REGION Network 3: Ya buscó caja DESACTIVADO
   // Detecta cuando el brazo de succion se encuentra arriba y setea una marca "ya buscó caja". La cinta no va a arrancar hasta que esta marca YA BUSCO CAJA se active.
   RUNG wire#powerrail
      Contact( "Marcha" )
      Contact( "iSNS_bs_arriba" )
      I_Contact( "iSNS_bs_abajo" )
      S_SR(operand := "Aux1", r1 := wire#w1)
      Coil( "Ya buscó caja" )
   END_RUNG
   RUNG wire#powerrail
      I_Contact( "Marcha" )
   END_RUNG wire#w1
   RUNG wire#powerrail
      { S7_Templates := "SrcType := DInt" } GE_Contact(in1 := "Encoder", in2 := 20)
      { S7_Templates := "SrcType := DInt" } LT_Contact(in1 := "Encoder", in2 := 45)
   END_RUNG wire#w1
   RUNG wire#powerrail
      Contact( "Habilita modo Probar" )
   END_RUNG wire#w1
   // the same network as SCL:
   IF "Marcha" AND "iSNS_bs_arriba" AND NOT "iSNS_bs_abajo" THEN
       "Aux1" := TRUE;   // SR flip-flop
   END_IF;
   IF NOT "Marcha" OR (("Encoder" >= 20) AND ("Encoder" < 45)) OR "Habilita modo Probar" THEN
       "Aux1" := FALSE;
   END_IF;
   "Ya buscó caja" := "Aux1";
END_REGION

REGION Network 4: Activa los succionadores.
   "TOFF".TOF(IN := NOT "iSNS_bs_abajo", PT := T#300ms);
   "Activa succionadores" := "TOFF".Q;
END_REGION

REGION Network 5: Cuando el brazo llega hasta abajo, lo detiene por 300 ms para asegurar que la caja salió de su rango. DESACTIVADO
   // DESACTIVADO
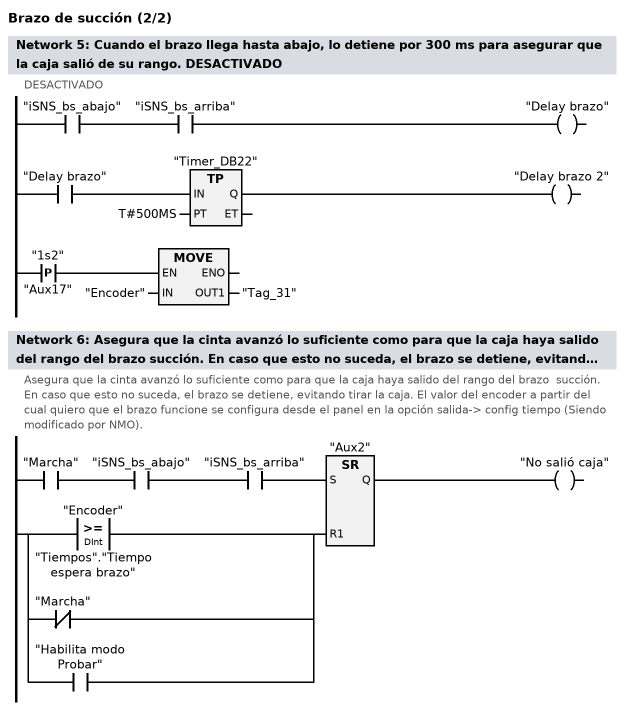
   "Delay brazo" := "iSNS_bs_abajo" AND "iSNS_bs_arriba";
   "Timer_DB22".TP(IN := "Delay brazo", PT := T#500MS);
   "Delay brazo 2" := "Timer_DB22".Q;
   #_w1 := "1s2" AND NOT "Aux17";   // rising edge of "1s2"
   "Aux17" := "1s2";
   IF #_w1 THEN "Tag_31" := "Encoder"; END_IF;
END_REGION

REGION Network 6: Asegura que la cinta avanzó lo suficiente como para que la caja haya salido del rango del brazo succión. En caso que esto no suceda, el brazo se detiene, evitando tirar la caja
   // Asegura que la cinta avanzó lo suficiente como para que la caja haya salido del rango del brazo  succión. En caso que esto no suceda, el brazo se detiene, evitando tirar la caja. El valor del encoder a partir del cual quiero que el brazo funcione se configura desde el panel en la opción salida-> config tiempo (Siendo modificado por NMO).
   RUNG wire#powerrail
      Contact( "Marcha" )
      Contact( "iSNS_bs_abajo" )
      Contact( "iSNS_bs_arriba" )
      S_SR(operand := "Aux2", r1 := wire#w1)
      Coil( "No salió caja" )
   END_RUNG
   RUNG wire#powerrail
      { S7_Templates := "SrcType := DInt" } GE_Contact(in1 := "Encoder", in2 := "Tiempos"."Tiempo espera brazo")
   END_RUNG wire#w1
   RUNG wire#powerrail
      I_Contact( "Marcha" )
   END_RUNG wire#w1
   RUNG wire#powerrail
      Contact( "Habilita modo Probar" )
   END_RUNG wire#w1
   // the same network as SCL:
   IF "Marcha" AND "iSNS_bs_abajo" AND "iSNS_bs_arriba" THEN
       "Aux2" := TRUE;   // SR flip-flop
   END_IF;
   IF ("Encoder" >= "Tiempos"."Tiempo espera brazo") OR NOT "Marcha" OR "Habilita modo Probar" THEN
       "Aux2" := FALSE;
   END_IF;
   "No salió caja" := "Aux2";
END_REGION
END_FUNCTION

ORGANIZATION_BLOCK "Main"   // OB1, LAD, ProgramCycle
TITLE = "Main Program Sweep (Cycle)"
{ S7_Optimized_Access := 'TRUE' }
VERSION : 0.1
BEGIN

REGION Network 1: Inversión de algunas entradas
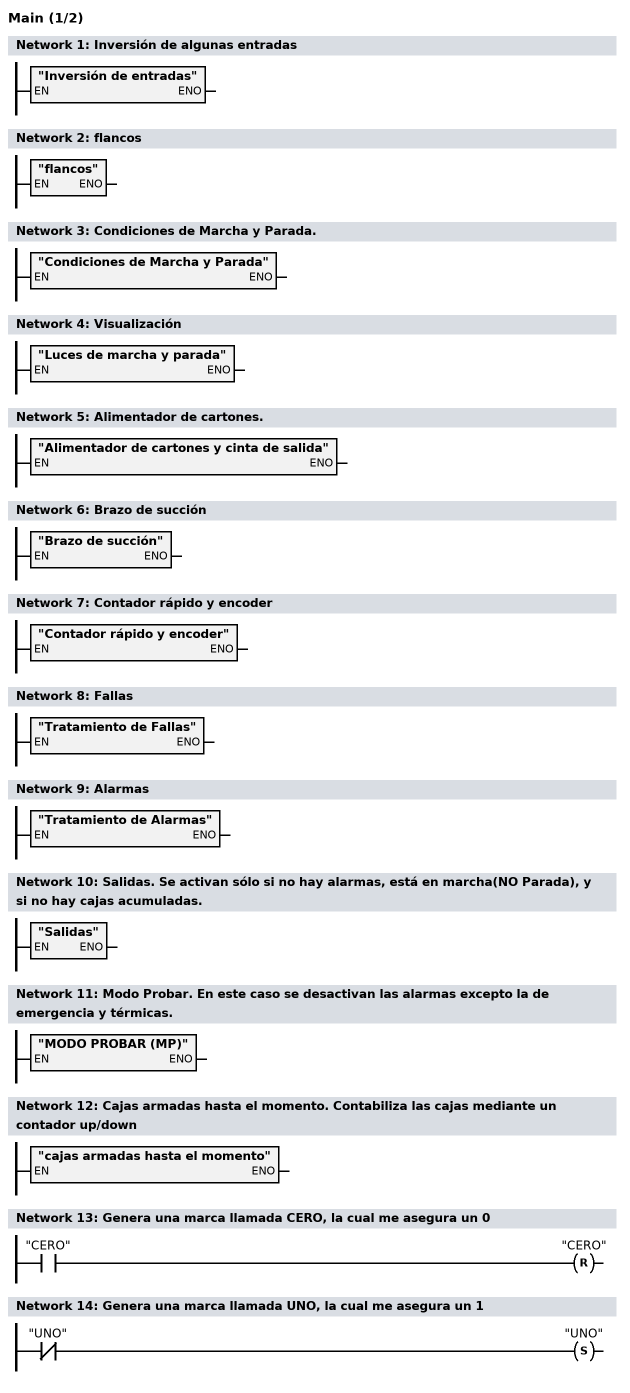
   RUNG wire#powerrail
      "Inversión de entradas"()
   END_RUNG
   // the same network as SCL:
   "Inversión de entradas"();
END_REGION

REGION Network 2: flancos
   RUNG wire#powerrail
      "flancos"()
   END_RUNG
   // the same network as SCL:
   "flancos"();
END_REGION

REGION Network 3: Condiciones de Marcha y Parada.
   RUNG wire#powerrail
      "Condiciones de Marcha y Parada"()
   END_RUNG
   // the same network as SCL:
   "Condiciones de Marcha y Parada"();
END_REGION

REGION Network 4: Visualización
   RUNG wire#powerrail
      "Luces de marcha y parada"()
   END_RUNG
   // the same network as SCL:
   "Luces de marcha y parada"();
END_REGION

REGION Network 5: Alimentador de cartones.
   RUNG wire#powerrail
      "Alimentador de cartones y cinta de salida"()
   END_RUNG
   // the same network as SCL:
   "Alimentador de cartones y cinta de salida"();
END_REGION

REGION Network 6: Brazo de succión
   RUNG wire#powerrail
      "Brazo de succión"()
   END_RUNG
   // the same network as SCL:
   "Brazo de succión"();
END_REGION

REGION Network 7: Contador rápido y encoder
   RUNG wire#powerrail
      "Contador rápido y encoder"()
   END_RUNG
   // the same network as SCL:
   "Contador rápido y encoder"();
END_REGION

REGION Network 8: Fallas
   RUNG wire#powerrail
      "Tratamiento de Fallas"()
   END_RUNG
   // the same network as SCL:
   "Tratamiento de Fallas"();
END_REGION

REGION Network 9: Alarmas
   RUNG wire#powerrail
      "Tratamiento de Alarmas"()
   END_RUNG
   // the same network as SCL:
   "Tratamiento de Alarmas"();
END_REGION

REGION Network 10: Salidas. Se activan sólo si no hay alarmas, está en marcha(NO Parada), y si no hay cajas acumuladas.
   RUNG wire#powerrail
      "Salidas"()
   END_RUNG
   // the same network as SCL:
   "Salidas"();
END_REGION

REGION Network 11: Modo Probar. En este caso se desactivan las alarmas excepto la de emergencia y térmicas.
   RUNG wire#powerrail
      "MODO PROBAR (MP)"()
   END_RUNG
   // the same network as SCL:
   "MODO PROBAR (MP)"();
END_REGION

REGION Network 12: Cajas armadas hasta el momento. Contabiliza las cajas mediante un contador up/down
   RUNG wire#powerrail
      "cajas armadas hasta el momento"()
   END_RUNG
   // the same network as SCL:
   "cajas armadas hasta el momento"();
END_REGION

REGION Network 13: Genera una marca llamada CERO, la cual me asegura un 0
   RUNG wire#powerrail
      Contact( "CERO" )
      R_Coil( "CERO" )
   END_RUNG
   // the same network as SCL:
   IF "CERO" THEN "CERO" := FALSE; END_IF;
END_REGION

REGION Network 14: Genera una marca llamada UNO, la cual me asegura un 1
   RUNG wire#powerrail
      I_Contact( "UNO" )
      S_Coil( "UNO" )
   END_RUNG
   // the same network as SCL:
   IF NOT "UNO" THEN "UNO" := TRUE; END_IF;
END_REGION

REGION Network 15: Secuencia Principal
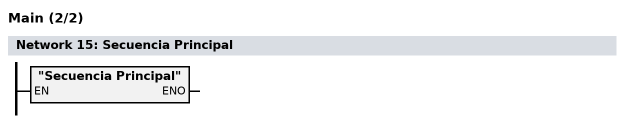
   RUNG wire#powerrail
      "Secuencia Principal"()
   END_RUNG
   // the same network as SCL:
   "Secuencia Principal"();
END_REGION
END_ORGANIZATION_BLOCK

(* ===== HMI "HMI_RT_1" =====
system functions are stored by id; their names below are inferred from use
connection "Conexión_HMI": ETHERNET, SMART_S7_1200_OMS

HMI tags "Tabla de variables estándar"
   "Alarmas_1" : Word AT %DB19.DBW0, 1 s
   "Alarmas_2" : Word AT %DB19.DBW2, 1 s
   "iAveria-reposicion" : Bool = PLC "iAveria-reposicion" AT %I32.2, 1 s
   "olmpR" : Bool = PLC oLmpR AT %Q32.5, 1 s
   "serie de fallas" : Bool = PLC "Serie de fallas" AT %M24.7, 1 s
   "Rearme desde panel" : Bool = PLC "Rearme desde panel" AT %M25.0, 1 s
   "olmpV" : Bool = PLC oLmpV AT %Q32.6, 1 s
   "SNS_carton en area de colado" : Bool = PLC "iSNS_carton en area de colado" AT %I33.3, 1 s
   "SNS_bs_arriba" : Bool = PLC iSNS_bs_arriba AT %I33.7, 1 s
   "SNS_bs_abajo" : Bool = PLC iSNS_bs_abajo AT %I33.6, 1 s
   "sns_nivel_bajo_cartones" : Bool = PLC iSNS_nivel_bajo_cartones AT %I33.0, 1 s
   "SNSpush_atras" : Bool = PLC iSNSpush_atras AT %I33.2, 1 s
   "SNSpush_adel" : Bool = PLC iSNSpush_adel AT %I0.2, 1 s
   "SNSpegamento en depósito" : Bool = PLC "iSNSpegamento en depósito" AT %I1.2, 1 s
   "SNScaja_trab" : Bool = PLC iSNScaja_trab AT %I1.4, 1 s
   "SNSalp" : Bool = PLC iSNSalp AT %I1.0, 1 s
   "SNScajas_acumuladas" : Bool = PLC iSnsCajaCerrada AT %I1.5, 1 s
   "om_cinta_principal" : Bool = PLC oM_cinta_principal AT %Q32.0, 1 s
   "om_bomba" : Bool = PLC oM_bomba AT %Q32.1, 1 s
   "oencola" : Bool = PLC oBoquilla_Encoladora AT %Q33.4, 1 s
   "om_brazo_succ" : Bool = PLC oM_brazo_succión AT %Q32.2, 1 s
   "om_pusher" : Bool = PLC oM_pusher AT %Q32.3, 1 s
   "om_cinta_sal" : Bool = PLC oM_cinta_sal AT %Q32.4, 1 s
   "osucción" : Bool = PLC oVálvula_Succión AT %Q33.0, 1 s
   "oagarra_solapas" : Bool = PLC oAgarra_solapas AT %Q33.1, 1 s
   "ocierra_solapa" : Bool = PLC oCierra_solapa AT %Q33.2, 1 s
   "opinza" : Bool = PLC oPinza AT %Q33.6, 1 s
   "oretB" : Bool = PLC oRetB AT %Q33.3, 1 s
   "oretC" : Bool = PLC oRetC AT %Q33.7, 1 s
   "oalim_cart" : Bool = PLC oAlim_cart AT %Q0.0, 1 s
   "opusher_out" : Bool = PLC oPusher_out AT %Q33.5, 1 s
   "iemergencia" : Bool = PLC iEmergencia AT %I32.1, 1 s
   "Emergencia desde panel" : Bool = PLC "Emergencia desde panel" AT %M25.1, 1 s
   "valor del encoder" : DWord = PLC "Valor del encoder" AT %MD180, 100 ms
   "Marcha desde panel" : Bool = PLC "Marcha desde panel" AT %M25.3, 1 s
   "Parada desde panel" : Bool = PLC Parada AT %M25.2, 1 s
   "S_automat" : Bool = PLC iS_automat AT %I33.4, 1 s
   "S_Probar" : Bool = PLC iS_Probar AT %I33.5, 1 s
   "Modo Manual" : Bool = PLC "Modo Manual" AT %M25.4, 1 s
   "K_encol_on" : Bool = PLC iK_encol_on AT %I33.1, 1 s
   "Valor cantidad de cajas armadas" : DWord = PLC "Valor cantidad de cajas armadas" AT %MD120, 1 s
   "Almacena el valor encolado experimental" : DWord = PLC "Exp Almacena el valor encolado experimental" AT %MD170, 1 s
   "ifase0" : Bool = PLC iFase0 AT %I0.3, 1 s
   "MPbrazo de succión arriba" : Bool = PLC "MPbrazo de succión arriba" AT %M40.0, 1 s
   "MPbrazo de succión abajo" : Bool = PLC "MPbrazo de succión abajo" AT %M40.1, 1 s
   "MPbotón activar pusher" : Bool = PLC "MPbotón activar pusher" AT %M42.0, 1 s
   "MPbotón Agarra solapas" : Bool = PLC "MPbotón Agarra solapas" AT %M41.3, 1 s
   "MPbotón activar retenedores de caja" : Bool = PLC "MPbotón activar retenedores de caja" AT %M43.4, 1 s
   "MPbotón Avanzar cinta por tramos" : Bool = PLC "MPbotón Avanzar cinta por tramos" AT %M41.6, 1 s
   "MPbotón alimentador de cartones" : Bool = PLC "MPbotón alimentador de cartones" AT %M41.2, 1 s
   "MPbotón Cierra solapa" : Bool = PLC "MPbotón Cierra solapa" AT %M41.4, 1 s
   "MPAcomodar brazo de succión" : Bool = PLC "MPAcomodar brazo de succión" AT %M43.6, 1 s
   "MPActiva bomba de vacío" : Bool = PLC "MPActiva bomba de vacío" AT %M42.5, 1 s
   "MPbotón Activar encoladora" : Bool = PLC "MPbotón Activar encoladora" AT %M41.0, 1 s
   "MPbotón Avanzar cinta" : Bool = PLC "MPbotón Avanzar cinta" AT %M41.5, 1 s
   "MPboton Activar bomba de vacío" : Bool = PLC "MPboton Activar bomba de vacío" AT %M40.7, 1 s
   "Rearmar" : Bool = PLC Rearmar AT %M23.1, 1 s
   "serie de Alarmas" : Bool = PLC "Serie de Alarmas" AT %M24.3, 1 s
   "P" : Bool = PLC iP AT %I32.6, 1 s
   "Marcha" : Bool = PLC Marcha AT %M20.0, 1 s
   "marca de prueba fase 0" : Bool = PLC "Exp marca de prueba fase 0" AT %M26.2, 1 s
   "Cajas acumuladas en salida" : Bool = PLC "Cajas acumuladas en salida" AT %M24.0, 1 s
   "k_EXT" : Bool = PLC k_EXT AT %I1.1, 1 s
   "ienable" : Bool = PLC iEnable AT %I32.0, 1 s
   "olinea-emergencia" : Bool = PLC "oLinea-emergencia" AT %Q32.7, 1 s
   "opacker" : Bool = PLC oPacker AT %Q0.3, 1 s
   "1s1" : Bool = PLC 1s1 AT %M0.0, 1 s
   "1s2" : Bool = PLC 1s2 AT %M0.1, 1 s
   "1s3" : Bool = PLC 1s3 AT %M0.2, 1 s
   "1s4" : Bool = PLC 1s4 AT %M0.3, 1 s
   "1s5" : Bool = PLC 1s5 AT %M0.4, 1 s
   "1s6" : Bool = PLC 1s6 AT %M0.5, 1 s
   "1s7" : Bool = PLC 1s7 AT %M0.6, 1 s
   "2s1" : Bool = PLC 2s1 AT %M4.0, 1 s
   "2s2" : Bool = PLC 2s2 AT %M4.1, 1 s
   "2s3" : Bool = PLC 2s3 AT %M4.2, 1 s
   "2s4" : Bool = PLC 2s4 AT %M4.3, 1 s
   "2s5" : Bool = PLC 2s5 AT %M4.4, 1 s
   "2s6" : Bool = PLC 2s6 AT %M4.5, 1 s
   "boton activar fingers" : Bool = PLC "Boton activar fingers" AT %M26.4, 1 s
   "osep_fing" : Bool = PLC oSep_fing AT %Q0.4, 1 s
   "botón packer" : Bool = PLC "Botón packer" AT %M26.5, 1 s
   "oquick_out" : Bool = PLC oQuick_out AT %Q0.1, 1 s
   "boton quick out" : Bool = PLC "Boton quick out" AT %M26.6, 1 s
   "Valor del encoder para calc encolado" : DWord = PLC "Exp valor del encoder para calc encolado" AT %MD220, 1 s
   "marca aux id118" : Bool = PLC "Exp marca aux id118" AT %M22.5, 1 s
   "Pulsador modo manual" : Bool = PLC "Pulsador modo manual" AT %M22.6, 1 s
   "MPvalor actual del encoder" : DWord = PLC "MPvalor actual del encoder" AT %MD200, 1 s
   "Aviso de cinta descalibrada probar" : Bool = PLC "Aviso de cinta descalibrada probar" AT %M22.7, 1 s
   "1s8" : Bool = PLC 1s8 AT %M0.7, 1 s
   "1s9" : Bool = PLC 1s9 AT %M1.0, 1 s
   "SNScaja_acum" : Bool = PLC iSNScaja_acum AT %I0.4, 1 s
   "datos de encolado_selcaja1000/1500" : Bool = PLC "datos de encolado".selcaja1000/1500 AT %DB11.DBX32.0, 1 s
   "parar proceso" : Bool = PLC "Parar proceso" AT %M29.5, 1 s
   "MPActivar cilindro pusher" : Bool = PLC "MPActivar cilindro pusher" AT %M42.2, 1 s
   "MPboton cilindro push" : Bool = PLC "MPboton cilindro push" AT %M44.0, 1 s
   "datos de encolado_Iniciosol1cj1000" : DInt = PLC "datos de encolado".Iniciosol1cj1000 AT %DB11.DBD0, 1 s
   "datos de encolado_finsol1cj1000" : DInt = PLC "datos de encolado".finsol1cj1000 AT %DB11.DBD4, 1 s
   "datos de encolado_Iniciosol2cj1000" : DInt = PLC "datos de encolado".Iniciosol2cj1000 AT %DB11.DBD8, 1 s
   "datos de encolado_finsol2cj1000" : DInt = PLC "datos de encolado".finsol2cj1000 AT %DB11.DBD12, 1 s
   "datos de encolado_Iniciosol1cj1500" : DInt = PLC "datos de encolado".Iniciosol1cj1500 AT %DB11.DBD16, 1 s
   "datos de encolado_finsol1cj1500" : DInt = PLC "datos de encolado".finsol1cj1500 AT %DB11.DBD20, 1 s
   "datos de encolado_Iniciosol2cj1500" : DInt = PLC "datos de encolado".Iniciosol2cj1500 AT %DB11.DBD24, 1 s
   "datos de encolado_finsol2cj1500" : DInt = PLC "datos de encolado".finsol2cj1500 AT %DB11.DBD28, 1 s
   "Resetear cajas armadas" : Bool = PLC "Resetear cajas armadas" AT %M25.5, 1 s
   "Tiempos_Tiempo cierra sol" : DInt = PLC Tiempos."Tiempo cierra sol" AT %DB23.DBD0, 1 s
   "Tiempos_Tiempo espera brazo" : DInt = PLC Tiempos."Tiempo espera brazo" AT %DB23.DBD4, 1 s
   "Valor encoder pusher salida" : DWord = PLC "Valor encoder pusher salida" AT %MD350, 1 s
   "Tiempos_tiempo cajas acum" : DInt = PLC Tiempos."tiempo cajas acum" AT %DB23.DBD8, 1 s
   "Tag_33" : Bool = PLC desactivar AT %M50.0, 1 s
   "AjusteEncoder_Hab_Pusher" : DInt = PLC AjusteEncoder.Hab_Pusher, 1 s
   "AjusteEncoder_Dhab_Pusher" : DInt = PLC AjusteEncoder.Dhab_Pusher, 1 s
   "AjusteEncoder_Reset" : Bool = PLC AjusteEncoder.Reset, 1 s
   "AjusteEncoder_Reset_Val" : DInt = PLC AjusteEncoder.Reset_Val, 1 s
   "HMI_Hab. Falla caja trab." : Bool = PLC "HMI_Hab. Falla caja trab." AT %M100.2, 1 s
   "Hab_Falla_Caja_Caida" : Bool = PLC HMI_Hab_Falla_Caja_Caida AT %M20.3, 1 s

discrete alarms
   1: 'Parada de Emergencia', class Alarmas sin acuse, trigger "Alarmas_1" bit 10
   2: 'Térmicas Brazo de succión y Pusher', class Alarmas sin acuse, trigger "Alarmas_1" bit 9
   3: 'Térmicas vacío, motor ppal, encoladora', class Alarmas sin acuse, trigger "Alarmas_1" bit 8
   4: 'Protección de Torque', class Alarmas sin acuse, trigger "Alarmas_1" bit 11
   5: 'falla en rele cadena', class Alarmas sin acuse, trigger "Alarmas_1" bit 12
   6: 'Falla en sensor atras Pusher', class Alarmas sin acuse, trigger "Alarmas_1" bit 13
   7: 'Falla en sensor adelante Pusher', class Alarmas sin acuse, trigger "Alarmas_1" bit 14
   8: 'Sensor brazo de succión de arriba', class Alarmas sin acuse, trigger "Alarmas_1" bit 15
   9: 'Sensor brazo de succión abajo', class Alarmas sin acuse, trigger "Alarmas_1" bit 0
   10: 'Sensor Área libre de Pusher', class Alarmas sin acuse, trigger "Alarmas_1" bit 1
   11: 'Sensor Alim Autom cartones', class Alarmas sin acuse, trigger "Alarmas_1" bit 2
   12: 'Encoder', class Alarmas sin acuse, trigger "Alarmas_1" bit 3
   13: 'Caja trabada en sector de salida', class Alarmas sin acuse, trigger "Alarmas_1" bit 4
   14: 'Incongruencia en sensores Pusher', class Alarmas sin acuse, trigger "Alarmas_1" bit 5
   15: 'Programacion prioritarias 1', class Alarmas sin acuse, trigger "Alarmas_1" bit 6
   16: 'Programación Concatenadoras 1', class Alarmas sin acuse, trigger "Alarmas_1" bit 7
   17: 'Programacion prioritarias 2', class Alarmas sin acuse, trigger "Alarmas_2" bit 8
   18: 'Programación Concatenadoras 2', class Alarmas sin acuse, trigger "Alarmas_2" bit 9
   19: 'Sensor área de encolado', class Alarmas sin acuse, trigger "Alarmas_2" bit 10
   20: 'Sin pegamento en depósito', class Alarmas sin acuse, trigger "Alarmas_2" bit 11
   21: 'falla en rele cadena 2', class Alarmas sin acuse, trigger "Alarmas_2" bit 12
   22: 'Caja Cerrada en la cadena', class Alarmas sin acuse, trigger "Alarmas_2" bit 13

text list "Nombre_imagen_lista_texto": 1 'Imagen raíz'; 2 'Imágenes de sistema'; 3 'Tareas varias'; 4 'Administración de usuarios'

screen "Alarmas" 800x480, template "Plantilla_1"
   Softkey "Softkey_F3" at 214,429 size 72x51
      on KeyUp: ActivateScreen("General", 0)
   AlarmView "Visor de avisos_1" at 5,100 size 785x254
   Button "Botón_1" at 12,364 size 780x68; TextOff 'Reconocer Alarmas'; TextOn 'Reconocido'
      on Press: SetBit("Rearme desde panel")
      on Release: ResetBit("Rearme desde panel")
   TextField "Campo de texto_1" at 140,440 size 122x36; Text 'Text'
   TextField "Campo de texto_9" at 268,440 size 125x36; Text 'Text'
   TextField "Campo de texto_10" at 398,440 size 122x36; Text 'Text'
   TextField "Campo de texto_7" at 0,6 size 800x56; Text 'Alarmas'
   Softkey "Softkey_F1" at 14,429 size 72x51
      on KeyUp: ActivateScreen("Sensores", 0)
   Softkey "Softkey_F2" at 114,429 size 72x51
      on KeyUp: ActivateScreen("Salidas", 0)

screen "Sensores" 800x480, template "Plantilla_1"
   Softkey "Softkey_F2" at 114,429 size 72x51
      on KeyDown: ActivateScreen("Salidas", 0)
   GraphicIOField "PlotLight_Round_G_2" at 418,156 size 42x34; PictureOn "PilotLight_Round_GN_Off_256c"; PictureOff "PilotLight_Round_N_On_mono"
      ProcessValue <- "SNS_carton en area de colado"
   GraphicIOField "PlotLight_Round_G_1" at 58,154 size 42x34; PictureOn "PilotLight_Round_GN_Off_256c"; PictureOff "PilotLight_Round_N_On_mono"
      ProcessValue <- "SNS_bs_arriba"
   GraphicIOField "PlotLight_Round_G_3" at 58,192 size 42x34; PictureOn "PilotLight_Round_GN_Off_256c"; PictureOff "PilotLight_Round_N_On_mono"
      ProcessValue <- "SNS_bs_abajo"
   GraphicIOField "PlotLight_Round_G_4" at 58,228 size 42x34; PictureOn "PilotLight_Round_GN_Off_256c"; PictureOff "PilotLight_Round_N_On_mono"
      ProcessValue <- "sns_nivel_bajo_cartones"
   GraphicIOField "PlotLight_Round_G_5" at 58,266 size 42x34; PictureOn "PilotLight_Round_GN_Off_256c"; PictureOff "PilotLight_Round_N_On_mono"
      ProcessValue <- "SNSpush_atras"
   GraphicIOField "PlotLight_Round_G_6" at 58,306 size 42x30; PictureOn "PilotLight_Round_GN_Off_256c"; PictureOff "PilotLight_Round_N_On_mono"
      ProcessValue <- "SNSpush_adel"
   GraphicIOField "PlotLight_Round_G_8" at 418,192 size 42x34; PictureOn "PilotLight_Round_N_On_mono"; PictureOff "PilotLight_Round_GN_Off_256c"
      ProcessValue <- "SNScaja_trab"
   GraphicIOField "PlotLight_Round_G_9" at 418,228 size 42x34; PictureOn "PilotLight_Round_GN_Off_256c"; PictureOff "PilotLight_Round_N_On_mono"
      ProcessValue <- "SNSalp"
   TextField "Campo de texto_2" at 475,154 size 200x27; Text 'Área encolado-B4440'
   GraphicIOField "PlotLight_Round_G_10" at 418,264 size 42x34; PictureOn "PilotLight_Round_N_On_mono"; PictureOff "PilotLight_Round_GN_Off_256c"
      ProcessValue <- "SNScaja_acum"
   TextField "Campo de texto_3" at 115,154 size 197x27; Text 'Brazo Arriba - B4480'
   TextField "Campo de texto_4" at 112,192 size 191x27; Text 'Brazo abajo - B4470'
   TextField "Campo de texto_5" at 112,230 size 216x27; Text 'Nivel bajo cart - B4410'
   TextField "Campo de texto_6" at 112,268 size 179x27; Text 'Push atrás - B4430'
   TextField "Campo de texto_7" at 112,306 size 167x27; Text 'Push Adel- B4140'
   TextField "Campo de texto_9" at 475,192 size 177x27; Text 'Caja en sal -B4250'
   TextField "Campo de texto_10" at 475,228 size 179x27; Text 'Área libre - B4210'
   TextField "Campo de texto_11" at 475,264 size 205x27; Text 'Caja en cta sal-B4450'
   TextField "Campo de texto_1" at 0,6 size 800x56; Text 'Sensores'
   TextField "Campo de texto_8" at 140,440 size 122x36; Text 'Salidas'
   TextField "Campo de texto_12" at 268,440 size 125x36; Text 'Text'
   TextField "Campo de texto_13" at 398,440 size 122x36; Text 'Text'

screen "Salidas" 800x480, template "Plantilla_1"
   Softkey "Softkey_F2" at 114,429 size 72x51
      on KeyDown: ActivateScreen("Sensores", 0)
   GraphicIOField "PlotLight_Round_G_2" at 438,176 size 42x34; PictureOff "PilotLight_Round_N_On_mono"; PictureOn "PilotLight_Round_GN_Off_256c"
      ProcessValue <- "om_cinta_principal"
   GraphicIOField "PlotLight_Round_G_1" at 438,360 size 42x34; PictureOff "PilotLight_Round_N_On_mono"; PictureOn "PilotLight_Round_GN_Off_256c"
      ProcessValue <- "om_bomba"
   GraphicIOField "PlotLight_Round_G_3" at 62,140 size 42x34; PictureOff "PilotLight_Round_N_On_mono"; PictureOn "PilotLight_Round_GN_Off_256c"
      ProcessValue <- "oencola"
   GraphicIOField "PlotLight_Round_G_4" at 62,176 size 42x34; PictureOff "PilotLight_Round_N_On_mono"; PictureOn "PilotLight_Round_GN_Off_256c"
      ProcessValue <- "om_brazo_succ"
   GraphicIOField "PlotLight_Round_G_5" at 62,212 size 42x34; PictureOff "PilotLight_Round_N_On_mono"; PictureOn "PilotLight_Round_GN_Off_256c"
      ProcessValue <- "om_pusher"
   GraphicIOField "PlotLight_Round_G_6" at 62,252 size 42x30; PictureOff "PilotLight_Round_N_On_mono"; PictureOn "PilotLight_Round_GN_Off_256c"
      ProcessValue <- "om_cinta_sal"
   GraphicIOField "PlotLight_Round_G_7" at 62,286 size 42x34; PictureOff "PilotLight_Round_N_On_mono"; PictureOn "PilotLight_Round_GN_Off_256c"
      ProcessValue <- "osucción"
   GraphicIOField "PlotLight_Round_G_8" at 62,324 size 42x34; PictureOff "PilotLight_Round_N_On_mono"; PictureOn "PilotLight_Round_GN_Off_256c"
      ProcessValue <- "oagarra_solapas"
   GraphicIOField "PlotLight_Round_G_9" at 62,360 size 42x34; PictureOff "PilotLight_Round_N_On_mono"; PictureOn "PilotLight_Round_GN_Off_256c"
      ProcessValue <- "ocierra_solapa"
   TextField "Campo de texto_2" at 498,176 size 166x27; Text 'Cinta ppal- Q32.0'
   GraphicIOField "PlotLight_Round_G_10" at 438,140 size 42x34; PictureOff "PilotLight_Round_N_On_mono"; PictureOn "PilotLight_Round_GN_Off_256c"
      ProcessValue <- "opinza"
   TextField "Campo de texto_3" at 498,362 size 121x27; Text 'Vacío- Q32.1'
   TextField "Campo de texto_5" at 120,178 size 139x27; Text 'Brazo s- Q32.2'
   TextField "Campo de texto_6" at 120,214 size 135x27; Text 'Pusher- Q32.3'
   TextField "Campo de texto_7" at 120,252 size 151x27; Text 'Cinta sal- Q32.4'
   TextField "Campo de texto_8" at 120,288 size 143x27; Text 'Succión- Q33.0'
   TextField "Campo de texto_9" at 120,326 size 173x27; Text 'Agarra sol - Q33.1'
   TextField "Campo de texto_11" at 495,138 size 120x27; Text 'Pinza- Q33.6'
   GraphicIOField "PlotLight_Round_G_11" at 438,324 size 42x34; PictureOff "PilotLight_Round_N_On_mono"; PictureOn "PilotLight_Round_GN_Off_256c"
      ProcessValue <- "oretB"
   TextField "Campo de texto_12" at 498,326 size 122x27; Text 'Ret B- Q33.7'
   GraphicIOField "PlotLight_Round_G_12" at 438,212 size 42x34; PictureOff "PilotLight_Round_N_On_mono"; PictureOn "PilotLight_Round_GN_Off_256c"
      ProcessValue <- "oretC"
   TextField "Campo de texto_13" at 498,214 size 122x27; Text 'Ret C- Q33.3'
   GraphicIOField "PlotLight_Round_G_13" at 438,250 size 42x34; PictureOff "PilotLight_Round_N_On_mono"; PictureOn "PilotLight_Round_GN_Off_256c"
      ProcessValue <- "oalim_cart"
   TextField "Campo de texto_14" at 498,252 size 144x27; Text 'Alim cart- Q0.0'
   GraphicIOField "PlotLight_Round_G_14" at 438,286 size 42x34; PictureOff "PilotLight_Round_N_On_mono"; PictureOn "PilotLight_Round_GN_Off_256c"
      ProcessValue <- "opusher_out"
   TextField "Campo de texto_15" at 498,288 size 153x27; Text 'Push out- Q33.5'
   TextField "Campo de texto_16" at 120,138 size 187x27; Text 'Boq Encolad- Q33.4'
   TextField "Campo de texto_10" at 120,362 size 151x27; Text 'Cierra sol Q33.2'
   TextField "Campo de texto_4" at 140,440 size 122x36; Text 'Sensores'
   TextField "Campo de texto_17" at 268,440 size 125x36; Text 'Text'
   TextField "Campo de texto_18" at 398,440 size 122x36; Text 'Text'
   TextField "Campo de texto_1" at 0,6 size 800x56; Text 'Salidas'

screen "General" 800x480, template "Plantilla_1"
   Softkey "Softkey_F2" at 114,429 size 72x51
      on KeyDown: ActivateScreen("Config - 1", 0)
   Softkey "Softkey_F3" at 214,429 size 72x51
      on KeyDown: ActivateScreen("Estado Actual", 0)
   Softkey "Softkey_F4" at 314,429 size 72x51
      on KeyDown: ActivateScreen("Sensores", 0)
   TextField "Campo de texto_2" at 40,122 size 134x37; Text 'En Marcha'
      Visibility <- "Marcha"
   TextField "Campo de texto_5" at 300,122 size 146x37; Text 'Automático'
      Visibility <- "S_automat"
   TextField "Campo de texto_6" at 325,122 size 85x37; Text 'Probar'
      Visibility <- "S_Probar"
   IOField "Campo ES_1" at 132,386 size 162x30; FormatPattern 999999
      ProcessValue <- "valor del encoder"
   IOField "Campo ES_2" at 138,250 size 520x46; FormatPattern 999999; Unit   Cajas Acumuladas
      ProcessValue <- "Valor cantidad de cajas armadas"
   TextField "Campo de texto_1" at 158,212 size 356x35; Text 'Cajas Acumuladas en la salida'
      Visibility <- "Cajas acumuladas en salida"
   Button "Botón_1" at 585,114 size 190x60; TextOff 'Paso Manual'
      on Press: SetBit("Pulsador modo manual")
      on Release: ResetBit("Pulsador modo manual")
      Appearance <- "Modo Manual"
   Button "Botón_2" at 320,310 size 132x44; TextOff 'Reset'; TextOn 'Reset cuenta'
      on Press: SetBit("Resetear cajas armadas")
      on Release: ResetBit("Resetear cajas armadas")
   TextField "Campo de texto_4" at 28,386 size 78x27; Text 'Encóder'
   TextField "Campo de texto_7" at 148,440 size 115x36; Text 'Config.'
   TextField "Campo de texto_8" at 268,440 size 112x36; Text 'Estado'
   TextField "Campo de texto_9" at 385,440 size 138x36; Text 'Diagnóstico'
   TextField "Campo de texto_3" at 0,6 size 800x56; Text 'General'
   TextField "Campo de texto_10" at 40,122 size 117x37; Text 'Detenido'
      Visibility <- "Marcha"
   TextField "Campo de texto_11" at 329,124 size 93x37; Text 'Manual'
      Visibility <- "Modo Manual"

Template "Plantilla_1" 800x480
   Softkey "Softkey_F1" at 14,429 size 72x51
      on KeyUp: ActivateScreen("General", 0)
   Softkey "Softkey_F6" at 514,429 size 72x51
      on KeyUp: ActivateScreen("Alarmas", 0)
   Softkey "Softkey_F5" at 414,429 size 72x51
      on KeyUp: ActivateScreen("Modo Probar", 0)
   DateTimeField "Plantilla_Campo de fecha y hora_1" at 512,54 size 195x30
      ProcessValue <- "HSC_reloj.YEAR"
   GraphicView "Plantilla_Visor de gráficos_1" at 20,14 size 162x40; Picture "eProC logo Gris 4"
   TextField "Campo de texto_1" at 5,440 size 132x36; Text 'General'
   TextField "Campo de texto_3" at 655,440 size 138x36; Text 'Alarmas'
   TextField "Campo de texto_5" at 525,440 size 125x36; Text 'Probar'
   TextField "Plantilla_Campo de texto_1" at 20,54 size 122x27; Text 'e013001v043'

screen "Modo Probar" 800x480, template "Plantilla_1"
   Button "Botón_2" at 160,366 size 222x60; TextOff 'Cierra solapa'
      on Press: SetBit("MPbotón Cierra solapa")
      on Release: ResetBit("MPbotón Cierra solapa")
   Button "Botón_3" at 422,366 size 222x60; TextOff 'Agarra solapas'
      on Press: SetBit("MPbotón Agarra solapas")
      on Release: ResetBit("MPbotón Agarra solapas")
   Button "Botón_5" at 422,302 size 222x60; TextOff 'Pusher y pinza'
      on Click: SetBit("MPbotón activar pusher")
   Button "Botón_7" at 422,174 size 222x60; TextOff 'Colero'
      on Click: ActivateScreen("Colero", 0)
   Button "Botón_8" at 160,302 size 222x60; TextOff 'Vacío y Succ'
      on Press: SetBit("MPboton Activar bomba de vacío")
      on Release: ResetBit("MPboton Activar bomba de vacío")
   Button "Botón_11" at 422,238 size 222x60; TextOff 'Retenedores'
      on Press: SetBit("MPbotón activar retenedores de caja")
      on Release: ResetBit("MPbotón activar retenedores de caja")
   Button "Botón_13" at 422,110 size 222x60; TextOff 'Alim carton'
      on Press: SetBit("MPbotón alimentador de cartones")
      on Release: ResetBit("MPbotón alimentador de cartones")
   Button "Botón_15" at 160,110 size 222x60; TextOff 'Acomodar brazo'
      on Press: SetBit("MPAcomodar brazo de succión")
      on Release: ResetBit("MPAcomodar brazo de succión")
   Button "Botón_16" at 160,174 size 222x60; TextOff 'Acomodar Cinta'
      on Click: SetBit("MPbotón Avanzar cinta por tramos")
   IOField "Campo ES_1" at 60,186 size 78x38; FormatPattern 999
      ProcessValue <- "valor del encoder"
   Button "Botón_1" at 160,238 size 222x60; TextOff 'Cil push'
      on Press: SetBit("MPboton cilindro push")
      on Release: ResetBit("MPboton cilindro push")
   TextField "Campo de texto_7" at 0,6 size 800x56; Text 'Modo Probar'
   TextField "Campo de texto_1" at 140,440 size 122x36; Text 'Text'
   TextField "Campo de texto_9" at 268,440 size 125x36; Text 'Text'
   TextField "Campo de texto_10" at 398,440 size 122x36; Text 'Text'

screen "Estado Actual" 800x480, template "Plantilla_1"
   TextField "Campo de texto_1" at 95,156 size 163x27; Text 'Estado 1: Reposo'
   TextField "Campo de texto_2" at 95,194 size 184x27; Text 'Estado2: Cinta Ppal'
   TextField "Campo de texto_3" at 95,232 size 205x27; Text 'Estado3: Retenedores'
   TextField "Campo de texto_4" at 95,270 size 206x27; Text 'Estado4: Desac Cinta'
   TextField "Campo de texto_5" at 95,308 size 153x27; Text 'Estado5: Pusher'
   TextField "Campo de texto_6" at 95,346 size 231x27; Text 'Estado6: Cilindro Pusher'
   TextField "Campo de texto_7" at 470,156 size 215x27; Text 'Estado7: Desac Pusher'
   TextField "Campo de texto_8" at 470,194 size 228x27; Text 'Estado8:Desac C Pusher'
   TextField "Campo de texto_9" at 470,232 size 188x27; Text 'Estado9: Fin Pusher'
   GraphicIOField "PlotLight_Round_G_2" at 40,158 size 42x34; PictureOff "PilotLight_Round_N_On_mono"; PictureOn "PilotLight_Round_GN_Off_256c"
      ProcessValue <- "1s1"
   GraphicIOField "PlotLight_Round_G_1" at 40,196 size 42x34; PictureOff "PilotLight_Round_N_On_mono"; PictureOn "PilotLight_Round_GN_Off_256c"
      ProcessValue <- "1s2"
   GraphicIOField "PlotLight_Round_G_3" at 40,234 size 42x34; PictureOff "PilotLight_Round_N_On_mono"; PictureOn "PilotLight_Round_GN_Off_256c"
      ProcessValue <- "1s3"
   GraphicIOField "PlotLight_Round_G_4" at 40,272 size 42x34; PictureOff "PilotLight_Round_N_On_mono"; PictureOn "PilotLight_Round_GN_Off_256c"
      ProcessValue <- "1s4"
   GraphicIOField "PlotLight_Round_G_5" at 40,310 size 42x34; PictureOff "PilotLight_Round_N_On_mono"; PictureOn "PilotLight_Round_GN_Off_256c"
      ProcessValue <- "1s5"
   GraphicIOField "PlotLight_Round_G_6" at 40,348 size 42x34; PictureOff "PilotLight_Round_N_On_mono"; PictureOn "PilotLight_Round_GN_Off_256c"
      ProcessValue <- "1s6"
   GraphicIOField "PlotLight_Round_G_7" at 415,158 size 42x34; PictureOff "PilotLight_Round_N_On_mono"; PictureOn "PilotLight_Round_GN_Off_256c"
      ProcessValue <- "1s7"
   GraphicIOField "PlotLight_Round_G_8" at 415,196 size 42x34; PictureOff "PilotLight_Round_N_On_mono"; PictureOn "PilotLight_Round_GN_Off_256c"
      ProcessValue <- "1s8"
   GraphicIOField "PlotLight_Round_G_9" at 415,234 size 42x34; PictureOff "PilotLight_Round_N_On_mono"; PictureOn "PilotLight_Round_GN_Off_256c"
      ProcessValue <- "1s9"
   TextField "Campo de texto_10" at 0,6 size 800x56; Text 'Estado'
   TextField "Campo de texto_11" at 140,440 size 122x36; Text 'Text'
   TextField "Campo de texto_12" at 268,440 size 125x36; Text 'Text'
   TextField "Campo de texto_13" at 398,440 size 122x36; Text 'Text'

screen "Colero" 800x480, template "Plantilla_1"
   GraphicIOField "PlotLight_Round_G_13" at 65,194 size 42x34; PictureOff "PilotLight_Round_N_On_mono"; PictureOn "PilotLight_Round_GN_Off_256c"
      ProcessValue <- "SNSpegamento en depósito"
   TextField "Campo de texto_15" at 125,188 size 213x26; Text 'Pegamento en depósito'
   TextField "Campo de texto_3" at 125,240 size 156x26; Text 'Colero Encendido'
   GraphicIOField "PlotLight_Round_G_1" at 65,244 size 42x32; PictureOff "PilotLight_Round_N_On_mono"; PictureOn "PilotLight_Round_GN_Off_256c"
      ProcessValue <- "K_encol_on"
   GraphicIOField "PlotLight_Round_G_2" at 65,290 size 42x34; PictureOff "PilotLight_Round_N_On_mono"; PictureOn "PilotLight_Round_GN_Off_256c"
      ProcessValue <- "SNS_carton en area de colado"
   TextField "Campo de texto_2" at 125,290 size 222x26; Text 'Sensor área de encolado'
   GraphicIOField "PlotLight_Round_G_3" at 65,144 size 42x34; PictureOff "PilotLight_Round_N_On_mono"; PictureOn "PilotLight_Round_GN_Off_256c"
      ProcessValue <- "oencola"
   TextField "Campo de texto_16" at 125,144 size 177x26; Text 'Boquilla Encoladora'
   Button "Botón_7" at 502,346 size 232x60; TextOff 'Probar PICOS'
      on Release: ResetBit("MPbotón Activar encoladora")
      on Press: SetBit("MPbotón Activar encoladora")
   TextField "Campo de texto_8" at 140,440 size 122x36; Text 'Text'
   TextField "Campo de texto_9" at 268,440 size 125x36; Text 'Text'
   TextField "Campo de texto_10" at 398,440 size 122x36; Text 'Text'
   TextField "Campo de texto_4" at 0,6 size 800x56; Text 'Colero'

screen "Config - 3" 800x480, template "Plantilla_1"
   Softkey "Softkey_F2" at 114,429 size 72x51
      on KeyDown: ActivateScreen("Config - 1", 0)
   Softkey "Softkey_F3" at 214,429 size 72x51
      on KeyDown: ActivateScreen("Config - 2", 0)
   Softkey "Softkey_F4" at 314,429 size 72x51
      on KeyDown: ActivateScreen("Config - 3", 0)
   IOField "Campo ES_1" at 130,272 size 95x30; FormatPattern s999
      ProcessValue <- "datos de encolado_Iniciosol1cj1000"
   IOField "Campo ES_2" at 135,378 size 95x30; FormatPattern s999
      ProcessValue <- "datos de encolado_Iniciosol2cj1000"
   IOField "Campo ES_3" at 258,272 size 95x30; FormatPattern s999
      ProcessValue <- "datos de encolado_finsol1cj1000"
   IOField "Campo ES_4" at 260,380 size 95x30; FormatPattern s999
      ProcessValue <- "datos de encolado_finsol2cj1000"
   TextField "Campo de texto_2" at 135,238 size 53x27; Text 'Inicio'
   TextField "Campo de texto_3" at 132,346 size 53x27; Text 'Inicio'
   TextField "Campo de texto_4" at 265,236 size 30x27; Text 'Fin'
   TextField "Campo de texto_5" at 265,346 size 30x27; Text 'Fin'
   IOField "Campo ES_5" at 468,274 size 95x30; FormatPattern s999
      ProcessValue <- "datos de encolado_Iniciosol1cj1500"
   IOField "Campo ES_6" at 472,380 size 95x30; FormatPattern s999
      ProcessValue <- "datos de encolado_Iniciosol2cj1500"
   IOField "Campo ES_7" at 590,276 size 95x30; FormatPattern s999
      ProcessValue <- "datos de encolado_finsol1cj1500"
   IOField "Campo ES_8" at 592,382 size 95x30; FormatPattern s999
      ProcessValue <- "datos de encolado_finsol2cj1500"
   TextField "Campo de texto_7" at 472,236 size 53x27; Text 'Inicio'
   TextField "Campo de texto_8" at 470,346 size 53x27; Text 'Inicio'
   TextField "Campo de texto_9" at 598,236 size 30x27; Text 'Fin'
   TextField "Campo de texto_10" at 598,346 size 30x27; Text 'Fin'
   TextField "Campo de texto_11" at 170,158 size 129x31; Text 'Cajas 1 litro'
   TextField "Campo de texto_12" at 480,154 size 160x31; Text 'Cajas 1.5 litros'
   TextField "Campo de texto_14" at 0,6 size 800x56; Text 'Referencias para Encolado'
   TextField "Campo de texto_1" at 135,204 size 82x27; Text 'Solapa 1'
   TextField "Campo de texto_6" at 132,312 size 82x27; Text 'Solapa 2'
   TextField "Campo de texto_13" at 475,204 size 82x27; Text 'Solapa 1'
   TextField "Campo de texto_15" at 472,312 size 82x27; Text 'Solapa 2'
   Switch "Interruptor_1" at 98,106 size 622x46; TextOff 'Cajas 1.5 Litro: Activado'; TextOn 'Cajas 1 litro: Activado'; CaptionText 'Switch'
      ProcessValue <- "datos de encolado_selcaja1000/1500"
   TextField "Campo de texto_16" at 140,440 size 122x36; Text 'Config 1'
   TextField "Campo de texto_17" at 268,440 size 125x36; Text 'Config 2'
   TextField "Campo de texto_18" at 398,440 size 122x36; Text 'Config 3'

screen "Config - 1" 800x480, template "Plantilla_1"
   Softkey "Softkey_F2" at 114,429 size 72x51
      on KeyDown: ActivateScreen("Config - 1", 0)
   Softkey "Softkey_F3" at 214,429 size 72x51
      on KeyDown: ActivateScreen("Config - 2", 0)
   Softkey "Softkey_F4" at 314,429 size 72x51
      on KeyDown: ActivateScreen("Config - 3", 0)
   IOField "Campo ES_1" at 272,124 size 85x30; FormatPattern 9999
      ProcessValue <- "Tiempos_Tiempo cierra sol"
   TextField "Campo de texto_1" at 32,120 size 181x27; Text 'Cierra solapa (ms)'
   TextField "Campo de texto_2" at 32,286 size 441x27; Text 'Referencia activación de brazo (70<valor<130)'
   IOField "Campo ES_2" at 40,334 size 92x32; FormatPattern s999
      ProcessValue <- "Tiempos_Tiempo espera brazo"
   TextField "Campo de texto_3" at 158,320 size 393x52; Text 'Valor de pulsos necesario para considerar que la caja salió del brazo de succión'
   TextField "Campo de texto_5" at 32,382 size 492x27; Text 'Valor = 0 indicaría que no se realiza ningún control'
   TextField "Campo de texto_4" at 35,160 size 366x77; Text 'Tiempo de retardo para desactivar el Cierra Solapa una véz que se activa la salida correspondiente'
   TextField "Campo de texto_7" at 0,6 size 800x56; Text 'Referencias Generales'
   TextField "Campo de texto_8" at 140,440 size 122x36; Text 'Config 1'
   TextField "Campo de texto_9" at 268,440 size 125x36; Text 'Config 2'
   TextField "Campo de texto_10" at 398,440 size 122x36; Text 'Config 3'

screen "Config - 2" 800x480, template "Plantilla_1"
   Softkey "Softkey_F2" at 114,429 size 72x51
      on KeyDown: ActivateScreen("Config - 1", 0)
   Softkey "Softkey_F3" at 214,429 size 72x51
      on KeyDown: ActivateScreen("Config - 2", 0)
   Softkey "Softkey_F4" at 314,429 size 72x51
      on KeyDown: ActivateScreen("Config - 3", 0)
   IOField "Campo ES_3" at 242,304 size 180x30; FormatPattern 9999; Unit  Pulsos
      ProcessValue <- "AjusteEncoder_Hab_Pusher"
   TextField "Campo de texto_7" at 68,254 size 170x27; Text 'Control de Pusher'
   IOField "Campo ES_4" at 242,344 size 180x30; FormatPattern 9999; Unit  Pulsos
      ProcessValue <- "AjusteEncoder_Dhab_Pusher"
   TextField "Campo de texto_8" at 48,340 size 142x27; Text 'Deshabilitación'
   IOField "Campo ES_2" at 70,136 size 165x38; FormatPattern 9999; Unit  Pulsos
      ProcessValue <- "AjusteEncoder_Reset_Val"
      Visibility <- "S_automat"
   TextField "Campo de texto_2" at 68,100 size 188x27; Text 'Forzado de Encóder'
   Button "Botón_1" at 250,134 size 150x44; TextOff 'Forzar'
      on Click: SetBit("AjusteEncoder_Reset")
      Visibility <- "S_automat"
   TextField "Campo de texto_14" at 0,6 size 800x56; Text 'Referencias para Pusher'
   TextField "Campo de texto_1" at 90,302 size 110x27; Text 'Habilitación'
   IOField "Campo ES_1" at 235,186 size 162x30; FormatPattern 999999
      ProcessValue <- "valor del encoder"
   TextField "Campo de texto_4" at 130,186 size 78x27; Text 'Encóder'
   TextField "Campo de texto_3" at 140,440 size 122x36; Text 'Config 1'
   TextField "Campo de texto_9" at 268,440 size 125x36; Text 'Config 2'
   TextField "Campo de texto_10" at 398,440 size 122x36; Text 'Config 3'
   Switch "Interruptor_1" at 565,322 size 160x64; TextOff 'OFF'; TextOn 'ON'; CaptionText 'Switch'
      ProcessValue <- "HMI_Hab. Falla caja trab."
   TextField "Campo de texto_5" at 532,258 size 173x52; Text 'activar/ desactivar falla caja trabada'
   Switch "Interruptor_2" at 565,178 size 160x64; TextOff 'OFF'; CaptionText 'Switch'; TextOn 'ON'
      ProcessValue <- "Hab_Falla_Caja_Caida"
   TextField "Campo de texto_6" at 525,116 size 173x52; Text 'activar/ desactivar falla caja cerrada'
*)